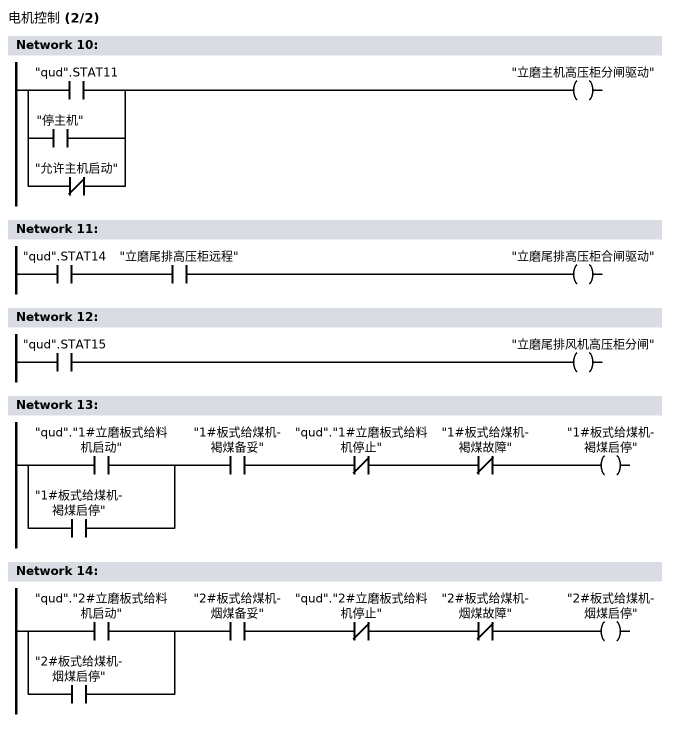
   RUNG wire#powerrail
      Contact( "qud".STAT11 )
      wire#w1
      Coil( "立磨主机高压柜分闸驱动" )
   END_RUNG
   RUNG wire#powerrail
      Contact( "停主机" )
   END_RUNG wire#w1
   RUNG wire#powerrail
      I_Contact( "允许主机启动" )
   END_RUNG wire#w1
   // the same network as SCL:
   "立磨主机高压柜分闸驱动" := "qud".STAT11 OR "停主机" OR NOT "允许主机启动";
END_REGION

REGION Network 11
   RUNG wire#powerrail
      Contact( "qud".STAT14 )
      Contact( "立磨尾排高压柜远程" )
      Coil( "立磨尾排高压柜合闸驱动" )
   END_RUNG
   // the same network as SCL:
   "立磨尾排高压柜合闸驱动" := "qud".STAT14 AND "立磨尾排高压柜远程";
END_REGION

REGION Network 12
   RUNG wire#powerrail
      Contact( "qud".STAT15 )
      Coil( "立磨尾排风机高压柜分闸" )
   END_RUNG
   // the same network as SCL:
   "立磨尾排风机高压柜分闸" := "qud".STAT15;
END_REGION

REGION Network 13
   RUNG wire#powerrail
      Contact( "qud"."1#立磨板式给料机启动" )
      wire#w1
      Contact( "1#板式给煤机-褐煤备妥" )
      I_Contact( "qud"."1#立磨板式给料机停止" )
      I_Contact( "1#板式给煤机-褐煤故障" )
      Coil( "1#板式给煤机-褐煤启停" )
   END_RUNG
   RUNG wire#powerrail
      Contact( "1#板式给煤机-褐煤启停" )
   END_RUNG wire#w1
   // the same network as SCL:
   "1#板式给煤机-褐煤启停" := ("qud"."1#立磨板式给料机启动" OR "1#板式给煤机-褐煤启停") AND "1#板式给煤机-褐煤备妥" AND NOT "qud"."1#立磨板式给料机停止" AND NOT "1#板式给煤机-褐煤故障";
END_REGION

REGION Network 14
   RUNG wire#powerrail
      Contact( "qud"."2#立磨板式给料机启动" )
      wire#w1
      Contact( "2#板式给煤机-烟煤备妥" )
      I_Contact( "qud"."2#立磨板式给料机停止" )
      I_Contact( "2#板式给煤机-烟煤故障" )
      Coil( "2#板式给煤机-烟煤启停" )
   END_RUNG
   RUNG wire#powerrail
      Contact( "2#板式给煤机-烟煤启停" )
   END_RUNG wire#w1
   // the same network as SCL:
   "2#板式给煤机-烟煤启停" := ("qud"."2#立磨板式给料机启动" OR "2#板式给煤机-烟煤启停") AND "2#板式给煤机-烟煤备妥" AND NOT "qud"."2#立磨板式给料机停止" AND NOT "2#板式给煤机-烟煤故障";
END_REGION
END_FUNCTION

FUNCTION "模拟量" : Void   // FC2, LAD
{ S7_Optimized_Access := 'FALSE' }
VERSION : 0.1
BEGIN

REGION Network 1
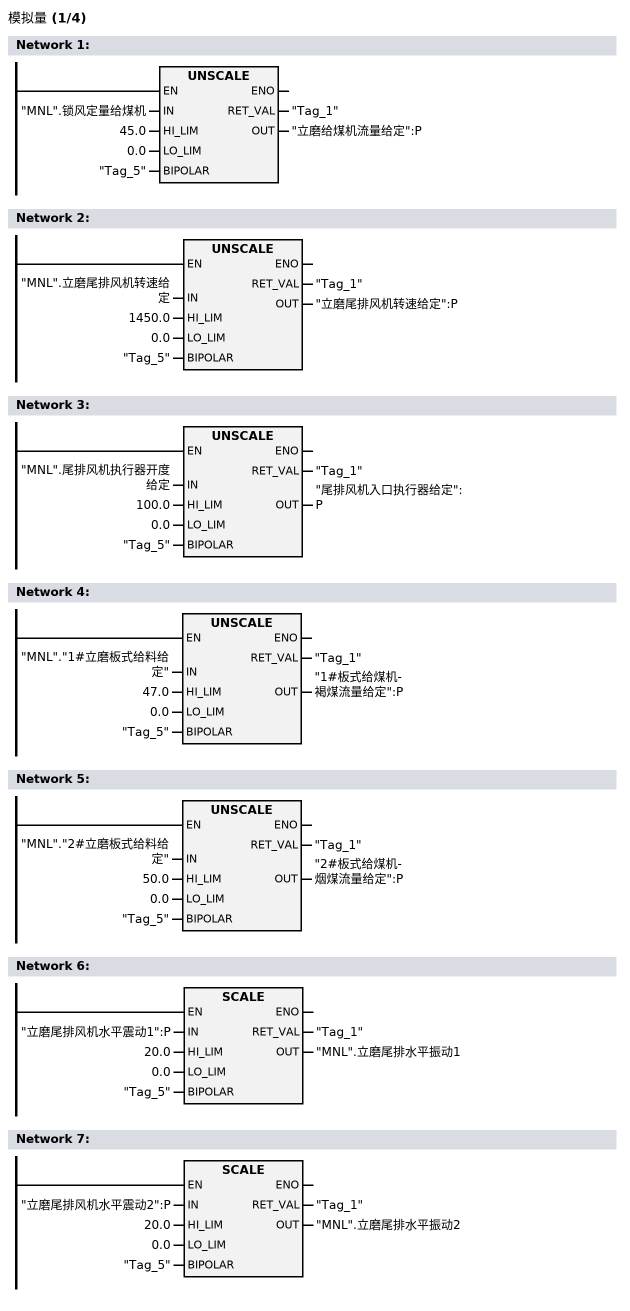
   "Tag_1" := UNSCALE(IN := "MNL".锁风定量给煤机,
                      HI_LIM := 45.0,
                      LO_LIM := 0.0,
                      BIPOLAR := "Tag_5",
                      OUT => "立磨给煤机流量给定":P);
END_REGION

REGION Network 2
   "Tag_1" := UNSCALE(IN := "MNL".立磨尾排风机转速给定,
                      HI_LIM := 1450.0,
                      LO_LIM := 0.0,
                      BIPOLAR := "Tag_5",
                      OUT => "立磨尾排风机转速给定":P);
END_REGION

REGION Network 3
   "Tag_1" := UNSCALE(IN := "MNL".尾排风机执行器开度给定,
                      HI_LIM := 100.0,
                      LO_LIM := 0.0,
                      BIPOLAR := "Tag_5",
                      OUT => "尾排风机入口执行器给定":P);
END_REGION

REGION Network 4
   "Tag_1" := UNSCALE(IN := "MNL"."1#立磨板式给料给定",
                      HI_LIM := 47.0,
                      LO_LIM := 0.0,
                      BIPOLAR := "Tag_5",
                      OUT => "1#板式给煤机-褐煤流量给定":P);
END_REGION

REGION Network 5
   "Tag_1" := UNSCALE(IN := "MNL"."2#立磨板式给料给定",
                      HI_LIM := 50.0,
                      LO_LIM := 0.0,
                      BIPOLAR := "Tag_5",
                      OUT => "2#板式给煤机-烟煤流量给定":P);
END_REGION

REGION Network 6
   "Tag_1" := SCALE(IN := "立磨尾排风机水平震动1":P,
                    HI_LIM := 20.0,
                    LO_LIM := 0.0,
                    BIPOLAR := "Tag_5",
                    OUT => "MNL".立磨尾排水平振动1);
END_REGION

REGION Network 7
   "Tag_1" := SCALE(IN := "立磨尾排风机水平震动2":P,
                    HI_LIM := 20.0,
                    LO_LIM := 0.0,
                    BIPOLAR := "Tag_5",
                    OUT => "MNL".立磨尾排水平振动2);
END_REGION

REGION Network 8
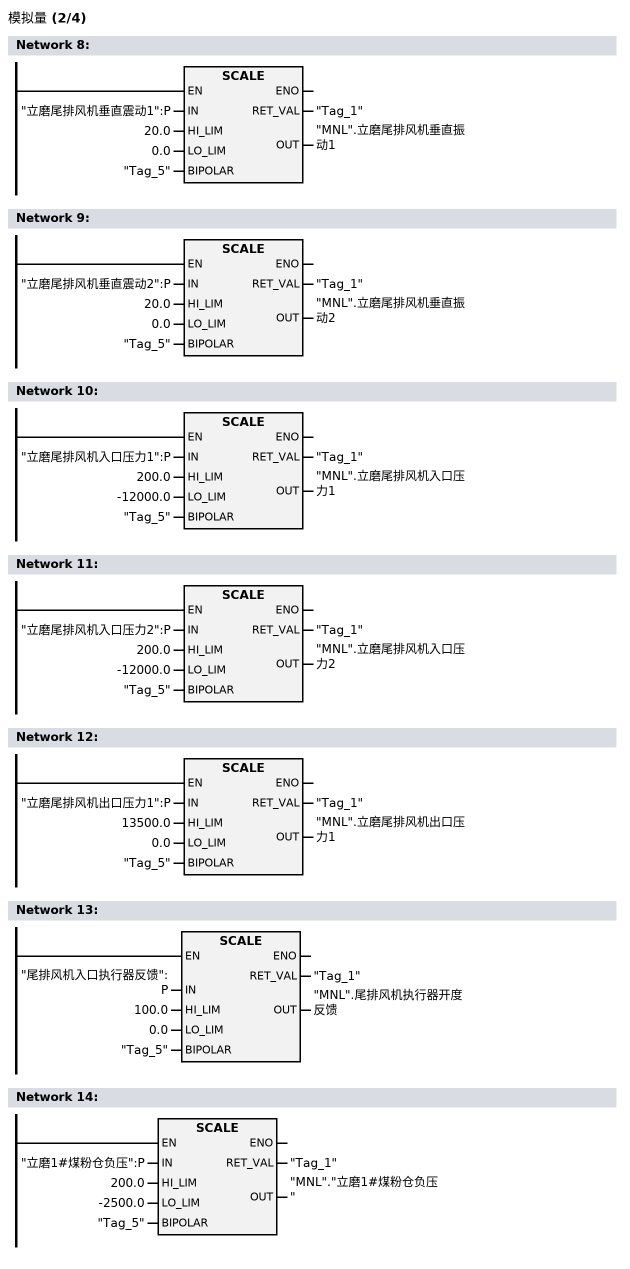
   "Tag_1" := SCALE(IN := "立磨尾排风机垂直震动1":P,
                    HI_LIM := 20.0,
                    LO_LIM := 0.0,
                    BIPOLAR := "Tag_5",
                    OUT => "MNL".立磨尾排风机垂直振动1);
END_REGION

REGION Network 9
   "Tag_1" := SCALE(IN := "立磨尾排风机垂直震动2":P,
                    HI_LIM := 20.0,
                    LO_LIM := 0.0,
                    BIPOLAR := "Tag_5",
                    OUT => "MNL".立磨尾排风机垂直振动2);
END_REGION

REGION Network 10
   "Tag_1" := SCALE(IN := "立磨尾排风机入口压力1":P,
                    HI_LIM := 200.0,
                    LO_LIM := -12000.0,
                    BIPOLAR := "Tag_5",
                    OUT => "MNL".立磨尾排风机入口压力1);
END_REGION

REGION Network 11
   "Tag_1" := SCALE(IN := "立磨尾排风机入口压力2":P,
                    HI_LIM := 200.0,
                    LO_LIM := -12000.0,
                    BIPOLAR := "Tag_5",
                    OUT => "MNL".立磨尾排风机入口压力2);
END_REGION

REGION Network 12
   "Tag_1" := SCALE(IN := "立磨尾排风机出口压力1":P,
                    HI_LIM := 13500.0,
                    LO_LIM := 0.0,
                    BIPOLAR := "Tag_5",
                    OUT => "MNL".立磨尾排风机出口压力1);
END_REGION

REGION Network 13
   "Tag_1" := SCALE(IN := "尾排风机入口执行器反馈":P,
                    HI_LIM := 100.0,
                    LO_LIM := 0.0,
                    BIPOLAR := "Tag_5",
                    OUT => "MNL".尾排风机执行器开度反馈);
END_REGION

REGION Network 14
   "Tag_1" := SCALE(IN := "立磨1#煤粉仓负压":P,
                    HI_LIM := 200.0,
                    LO_LIM := -2500.0,
                    BIPOLAR := "Tag_5",
                    OUT => "MNL"."立磨1#煤粉仓负压");
END_REGION

REGION Network 15
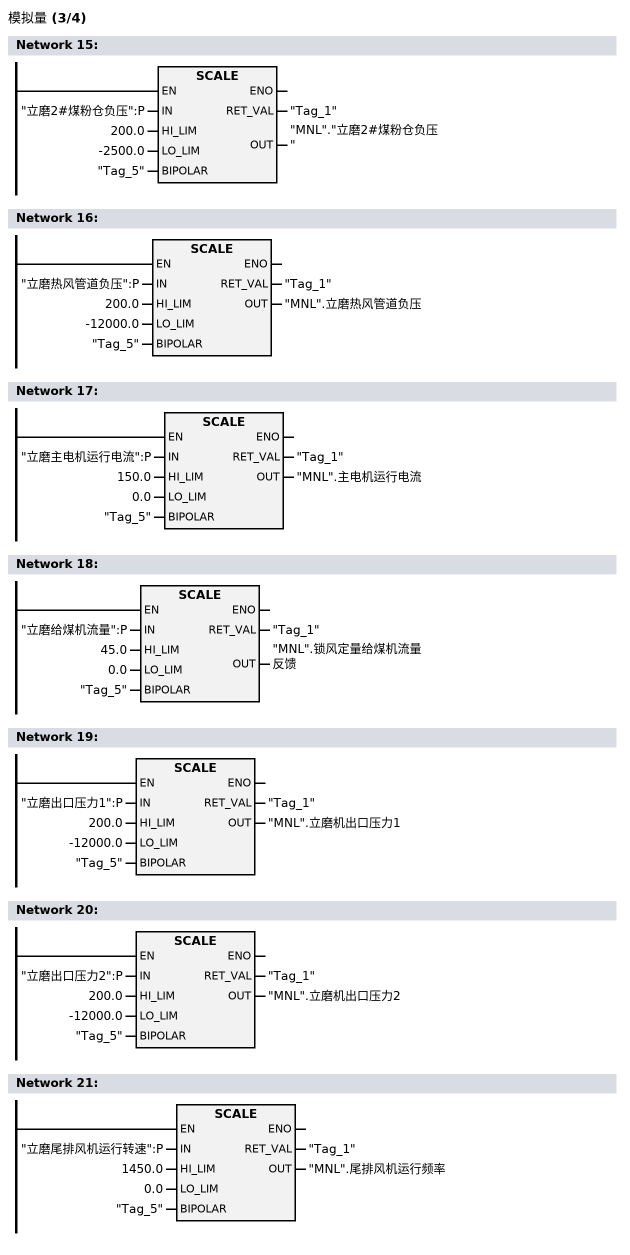
   "Tag_1" := SCALE(IN := "立磨2#煤粉仓负压":P,
                    HI_LIM := 200.0,
                    LO_LIM := -2500.0,
                    BIPOLAR := "Tag_5",
                    OUT => "MNL"."立磨2#煤粉仓负压");
END_REGION

REGION Network 16
   "Tag_1" := SCALE(IN := "立磨热风管道负压":P,
                    HI_LIM := 200.0,
                    LO_LIM := -12000.0,
                    BIPOLAR := "Tag_5",
                    OUT => "MNL".立磨热风管道负压);
END_REGION

REGION Network 17
   "Tag_1" := SCALE(IN := "立磨主电机运行电流":P,
                    HI_LIM := 150.0,
                    LO_LIM := 0.0,
                    BIPOLAR := "Tag_5",
                    OUT => "MNL".主电机运行电流);
END_REGION

REGION Network 18
   "Tag_1" := SCALE(IN := "立磨给煤机流量":P,
                    HI_LIM := 45.0,
                    LO_LIM := 0.0,
                    BIPOLAR := "Tag_5",
                    OUT => "MNL".锁风定量给煤机流量反馈);
END_REGION

REGION Network 19
   "Tag_1" := SCALE(IN := "立磨出口压力1":P,
                    HI_LIM := 200.0,
                    LO_LIM := -12000.0,
                    BIPOLAR := "Tag_5",
                    OUT => "MNL".立磨机出口压力1);
END_REGION

REGION Network 20
   "Tag_1" := SCALE(IN := "立磨出口压力2":P,
                    HI_LIM := 200.0,
                    LO_LIM := -12000.0,
                    BIPOLAR := "Tag_5",
                    OUT => "MNL".立磨机出口压力2);
END_REGION

REGION Network 21
   "Tag_1" := SCALE(IN := "立磨尾排风机运行转速":P,
                    HI_LIM := 1450.0,
                    LO_LIM := 0.0,
                    BIPOLAR := "Tag_5",
                    OUT => "MNL".尾排风机运行频率);
END_REGION

REGION Network 22
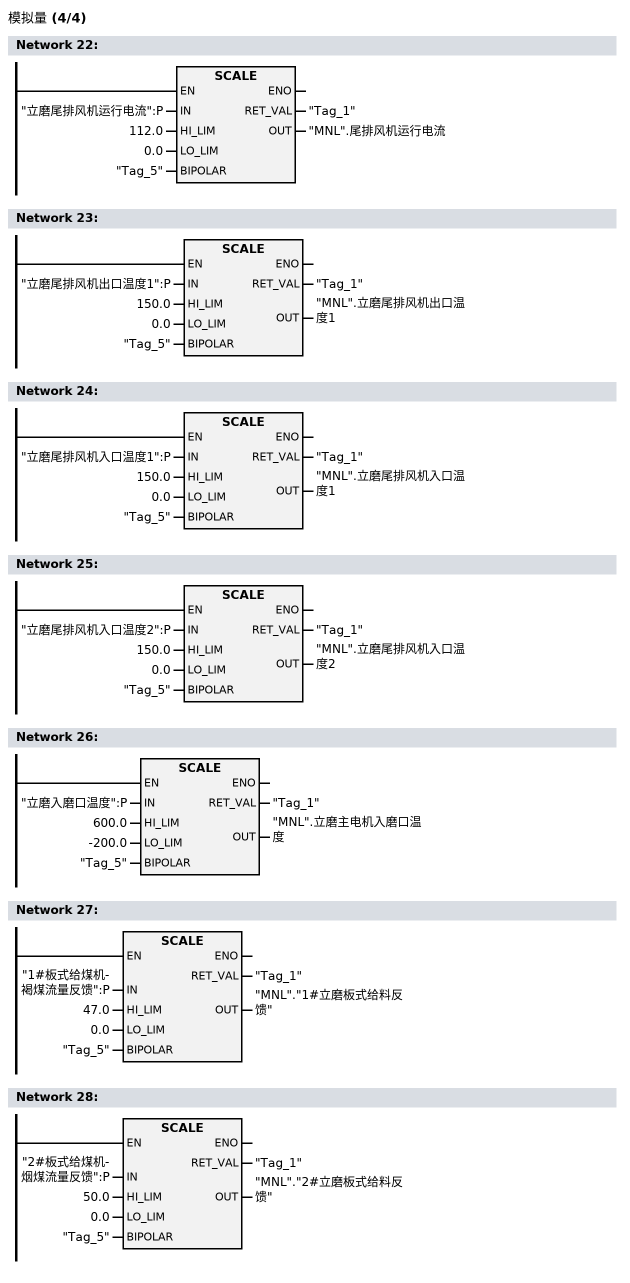
   "Tag_1" := SCALE(IN := "立磨尾排风机运行电流":P,
                    HI_LIM := 112.0,
                    LO_LIM := 0.0,
                    BIPOLAR := "Tag_5",
                    OUT => "MNL".尾排风机运行电流);
END_REGION

REGION Network 23
   "Tag_1" := SCALE(IN := "立磨尾排风机出口温度1":P,
                    HI_LIM := 150.0,
                    LO_LIM := 0.0,
                    BIPOLAR := "Tag_5",
                    OUT => "MNL".立磨尾排风机出口温度1);
END_REGION

REGION Network 24
   "Tag_1" := SCALE(IN := "立磨尾排风机入口温度1":P,
                    HI_LIM := 150.0,
                    LO_LIM := 0.0,
                    BIPOLAR := "Tag_5",
                    OUT => "MNL".立磨尾排风机入口温度1);
END_REGION

REGION Network 25
   "Tag_1" := SCALE(IN := "立磨尾排风机入口温度2":P,
                    HI_LIM := 150.0,
                    LO_LIM := 0.0,
                    BIPOLAR := "Tag_5",
                    OUT => "MNL".立磨尾排风机入口温度2);
END_REGION

REGION Network 26
   "Tag_1" := SCALE(IN := "立磨入磨口温度":P,
                    HI_LIM := 600.0,
                    LO_LIM := -200.0,
                    BIPOLAR := "Tag_5",
                    OUT => "MNL".立磨主电机入磨口温度);
END_REGION

REGION Network 27
   "Tag_1" := SCALE(IN := "1#板式给煤机-褐煤流量反馈":P,
                    HI_LIM := 47.0,
                    LO_LIM := 0.0,
                    BIPOLAR := "Tag_5",
                    OUT => "MNL"."1#立磨板式给料反馈");
END_REGION

REGION Network 28
   "Tag_1" := SCALE(IN := "2#板式给煤机-烟煤流量反馈":P,
                    HI_LIM := 50.0,
                    LO_LIM := 0.0,
                    BIPOLAR := "Tag_5",
                    OUT => "MNL"."2#立磨板式给料反馈");
END_REGION
END_FUNCTION

FUNCTION "料仓控制" : Void   // FC3, LAD
{ S7_Optimized_Access := 'FALSE' }
VERSION : 0.1
BEGIN

REGION Network 1
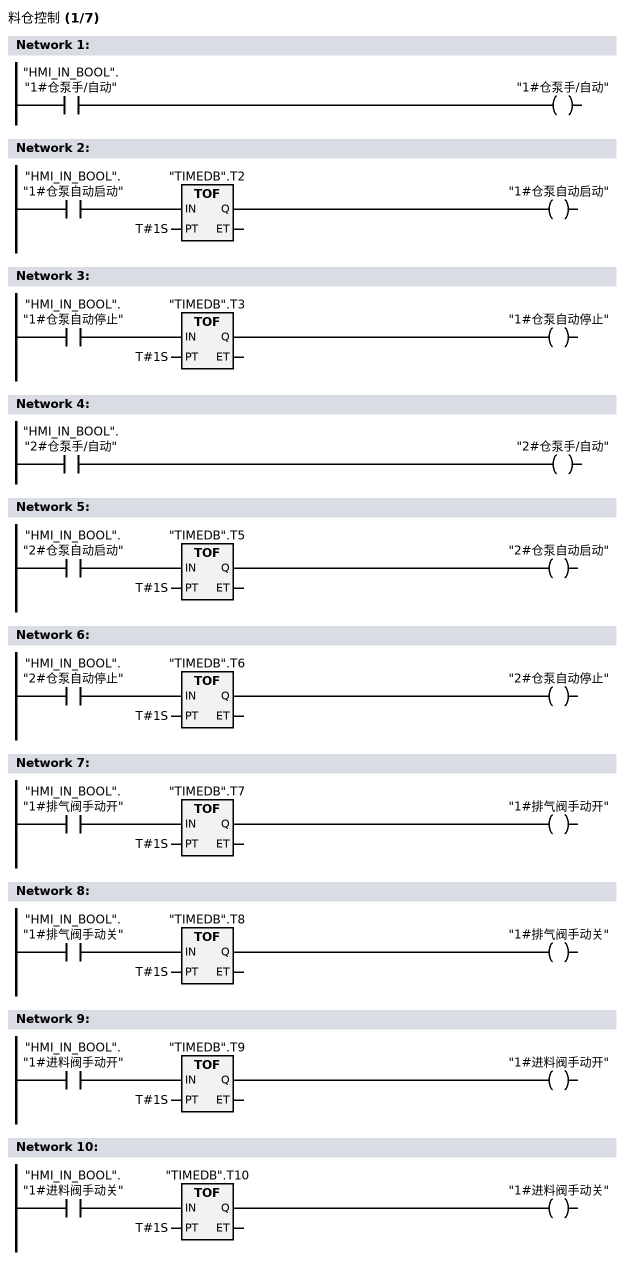
   RUNG wire#powerrail
      Contact( "HMI_IN_BOOL"."1#仓泵手/自动" )
      Coil( "1#仓泵手/自动" )
   END_RUNG
   // the same network as SCL:
   "1#仓泵手/自动" := "HMI_IN_BOOL"."1#仓泵手/自动";
END_REGION

REGION Network 2
   "TIMEDB".T2.TOF(IN := "HMI_IN_BOOL"."1#仓泵自动启动", PT := T#1S);
   "1#仓泵自动启动" := "TIMEDB".T2.Q;
END_REGION

REGION Network 3
   "TIMEDB".T3.TOF(IN := "HMI_IN_BOOL"."1#仓泵自动停止", PT := T#1S);
   "1#仓泵自动停止" := "TIMEDB".T3.Q;
END_REGION

REGION Network 4
   RUNG wire#powerrail
      Contact( "HMI_IN_BOOL"."2#仓泵手/自动" )
      Coil( "2#仓泵手/自动" )
   END_RUNG
   // the same network as SCL:
   "2#仓泵手/自动" := "HMI_IN_BOOL"."2#仓泵手/自动";
END_REGION

REGION Network 5
   "TIMEDB".T5.TOF(IN := "HMI_IN_BOOL"."2#仓泵自动启动", PT := T#1S);
   "2#仓泵自动启动" := "TIMEDB".T5.Q;
END_REGION

REGION Network 6
   "TIMEDB".T6.TOF(IN := "HMI_IN_BOOL"."2#仓泵自动停止", PT := T#1S);
   "2#仓泵自动停止" := "TIMEDB".T6.Q;
END_REGION

REGION Network 7
   "TIMEDB".T7.TOF(IN := "HMI_IN_BOOL"."1#排气阀手动开", PT := T#1S);
   "1#排气阀手动开" := "TIMEDB".T7.Q;
END_REGION

REGION Network 8
   "TIMEDB".T8.TOF(IN := "HMI_IN_BOOL"."1#排气阀手动关", PT := T#1S);
   "1#排气阀手动关" := "TIMEDB".T8.Q;
END_REGION

REGION Network 9
   "TIMEDB".T9.TOF(IN := "HMI_IN_BOOL"."1#进料阀手动开", PT := T#1S);
   "1#进料阀手动开" := "TIMEDB".T9.Q;
END_REGION

REGION Network 10
   "TIMEDB".T10.TOF(IN := "HMI_IN_BOOL"."1#进料阀手动关", PT := T#1S);
   "1#进料阀手动关" := "TIMEDB".T10.Q;
END_REGION

REGION Network 11
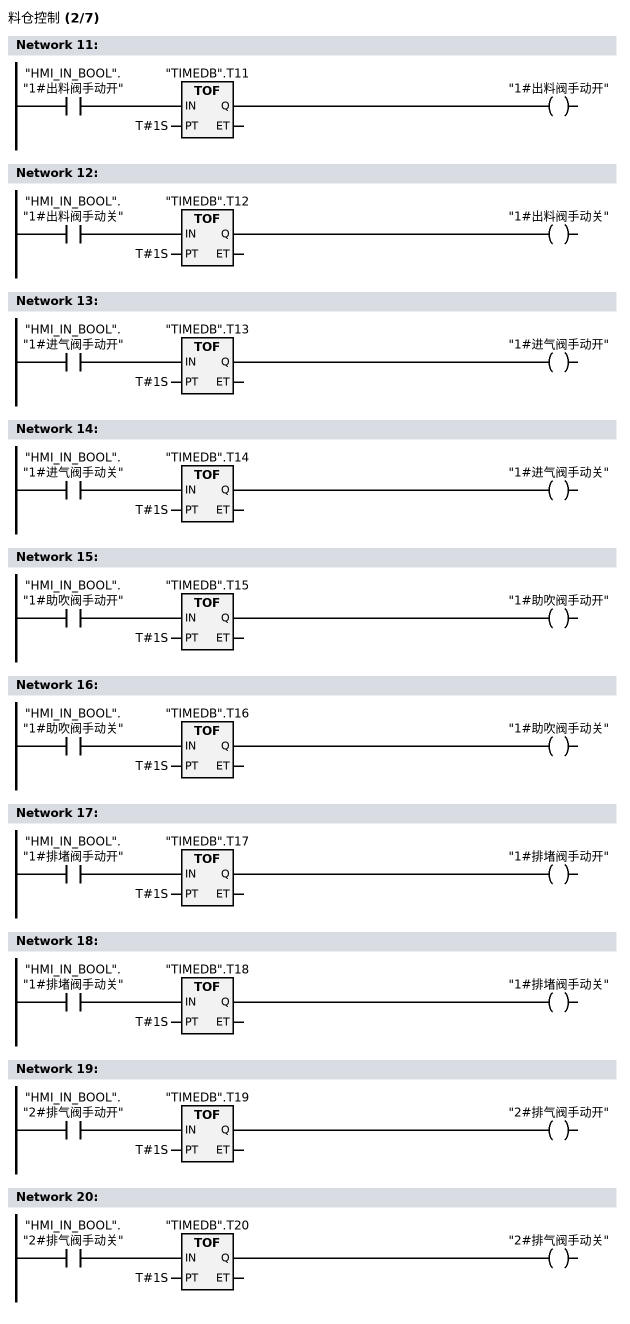
   "TIMEDB".T11.TOF(IN := "HMI_IN_BOOL"."1#出料阀手动开", PT := T#1S);
   "1#出料阀手动开" := "TIMEDB".T11.Q;
END_REGION

REGION Network 12
   "TIMEDB".T12.TOF(IN := "HMI_IN_BOOL"."1#出料阀手动关", PT := T#1S);
   "1#出料阀手动关" := "TIMEDB".T12.Q;
END_REGION

REGION Network 13
   "TIMEDB".T13.TOF(IN := "HMI_IN_BOOL"."1#进气阀手动开", PT := T#1S);
   "1#进气阀手动开" := "TIMEDB".T13.Q;
END_REGION

REGION Network 14
   "TIMEDB".T14.TOF(IN := "HMI_IN_BOOL"."1#进气阀手动关", PT := T#1S);
   "1#进气阀手动关" := "TIMEDB".T14.Q;
END_REGION

REGION Network 15
   "TIMEDB".T15.TOF(IN := "HMI_IN_BOOL"."1#助吹阀手动开", PT := T#1S);
   "1#助吹阀手动开" := "TIMEDB".T15.Q;
END_REGION

REGION Network 16
   "TIMEDB".T16.TOF(IN := "HMI_IN_BOOL"."1#助吹阀手动关", PT := T#1S);
   "1#助吹阀手动关" := "TIMEDB".T16.Q;
END_REGION

REGION Network 17
   "TIMEDB".T17.TOF(IN := "HMI_IN_BOOL"."1#排堵阀手动开", PT := T#1S);
   "1#排堵阀手动开" := "TIMEDB".T17.Q;
END_REGION

REGION Network 18
   "TIMEDB".T18.TOF(IN := "HMI_IN_BOOL"."1#排堵阀手动关", PT := T#1S);
   "1#排堵阀手动关" := "TIMEDB".T18.Q;
END_REGION

REGION Network 19
   "TIMEDB".T19.TOF(IN := "HMI_IN_BOOL"."2#排气阀手动开", PT := T#1S);
   "2#排气阀手动开" := "TIMEDB".T19.Q;
END_REGION

REGION Network 20
   "TIMEDB".T20.TOF(IN := "HMI_IN_BOOL"."2#排气阀手动关", PT := T#1S);
   "2#排气阀手动关" := "TIMEDB".T20.Q;
END_REGION

REGION Network 21
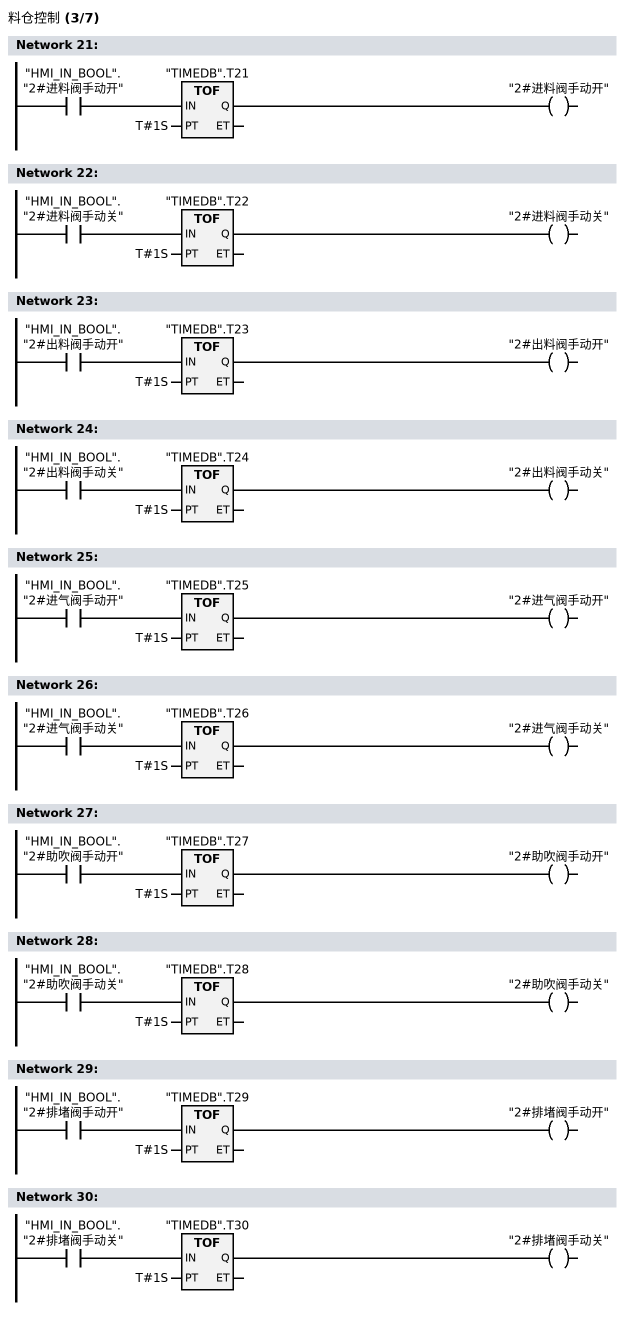
   "TIMEDB".T21.TOF(IN := "HMI_IN_BOOL"."2#进料阀手动开", PT := T#1S);
   "2#进料阀手动开" := "TIMEDB".T21.Q;
END_REGION

REGION Network 22
   "TIMEDB".T22.TOF(IN := "HMI_IN_BOOL"."2#进料阀手动关", PT := T#1S);
   "2#进料阀手动关" := "TIMEDB".T22.Q;
END_REGION

REGION Network 23
   "TIMEDB".T23.TOF(IN := "HMI_IN_BOOL"."2#出料阀手动开", PT := T#1S);
   "2#出料阀手动开" := "TIMEDB".T23.Q;
END_REGION

REGION Network 24
   "TIMEDB".T24.TOF(IN := "HMI_IN_BOOL"."2#出料阀手动关", PT := T#1S);
   "2#出料阀手动关" := "TIMEDB".T24.Q;
END_REGION

REGION Network 25
   "TIMEDB".T25.TOF(IN := "HMI_IN_BOOL"."2#进气阀手动开", PT := T#1S);
   "2#进气阀手动开" := "TIMEDB".T25.Q;
END_REGION

REGION Network 26
   "TIMEDB".T26.TOF(IN := "HMI_IN_BOOL"."2#进气阀手动关", PT := T#1S);
   "2#进气阀手动关" := "TIMEDB".T26.Q;
END_REGION

REGION Network 27
   "TIMEDB".T27.TOF(IN := "HMI_IN_BOOL"."2#助吹阀手动开", PT := T#1S);
   "2#助吹阀手动开" := "TIMEDB".T27.Q;
END_REGION

REGION Network 28
   "TIMEDB".T28.TOF(IN := "HMI_IN_BOOL"."2#助吹阀手动关", PT := T#1S);
   "2#助吹阀手动关" := "TIMEDB".T28.Q;
END_REGION

REGION Network 29
   "TIMEDB".T29.TOF(IN := "HMI_IN_BOOL"."2#排堵阀手动开", PT := T#1S);
   "2#排堵阀手动开" := "TIMEDB".T29.Q;
END_REGION

REGION Network 30
   "TIMEDB".T30.TOF(IN := "HMI_IN_BOOL"."2#排堵阀手动关", PT := T#1S);
   "2#排堵阀手动关" := "TIMEDB".T30.Q;
END_REGION

REGION Network 31
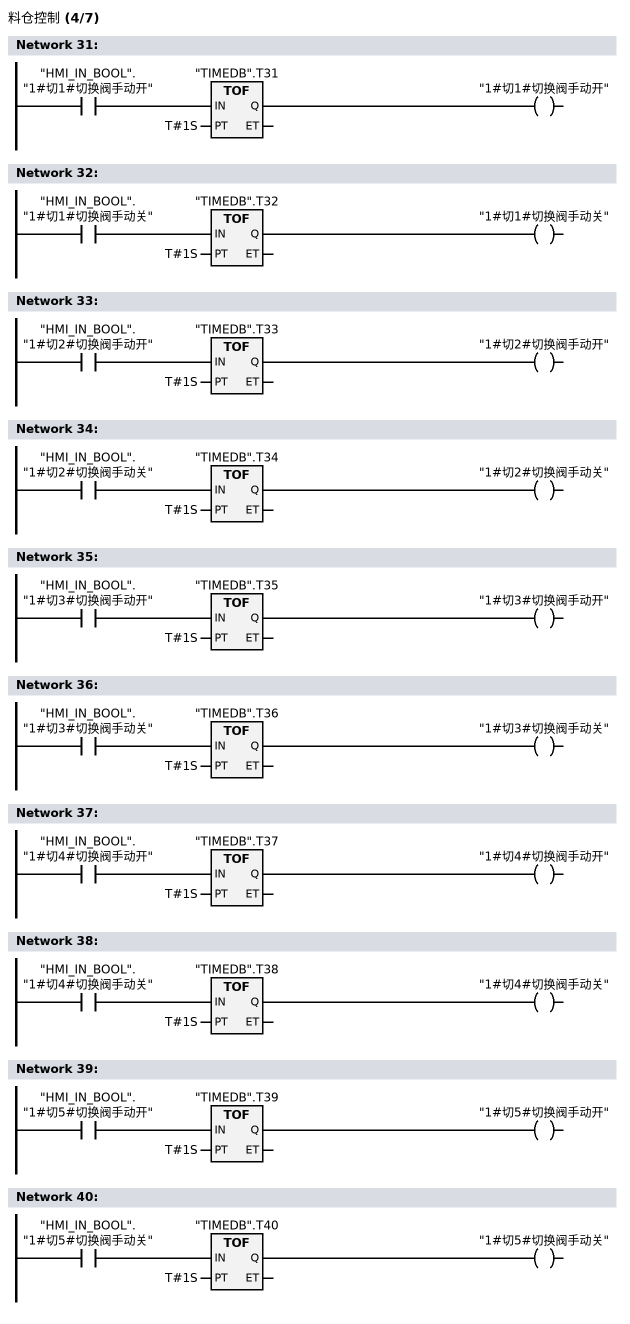
   "TIMEDB".T31.TOF(IN := "HMI_IN_BOOL"."1#切1#切换阀手动开", PT := T#1S);
   "1#切1#切换阀手动开" := "TIMEDB".T31.Q;
END_REGION

REGION Network 32
   "TIMEDB".T32.TOF(IN := "HMI_IN_BOOL"."1#切1#切换阀手动关", PT := T#1S);
   "1#切1#切换阀手动关" := "TIMEDB".T32.Q;
END_REGION

REGION Network 33
   "TIMEDB".T33.TOF(IN := "HMI_IN_BOOL"."1#切2#切换阀手动开", PT := T#1S);
   "1#切2#切换阀手动开" := "TIMEDB".T33.Q;
END_REGION

REGION Network 34
   "TIMEDB".T34.TOF(IN := "HMI_IN_BOOL"."1#切2#切换阀手动关", PT := T#1S);
   "1#切2#切换阀手动关" := "TIMEDB".T34.Q;
END_REGION

REGION Network 35
   "TIMEDB".T35.TOF(IN := "HMI_IN_BOOL"."1#切3#切换阀手动开", PT := T#1S);
   "1#切3#切换阀手动开" := "TIMEDB".T35.Q;
END_REGION

REGION Network 36
   "TIMEDB".T36.TOF(IN := "HMI_IN_BOOL"."1#切3#切换阀手动关", PT := T#1S);
   "1#切3#切换阀手动关" := "TIMEDB".T36.Q;
END_REGION

REGION Network 37
   "TIMEDB".T37.TOF(IN := "HMI_IN_BOOL"."1#切4#切换阀手动开", PT := T#1S);
   "1#切4#切换阀手动开" := "TIMEDB".T37.Q;
END_REGION

REGION Network 38
   "TIMEDB".T38.TOF(IN := "HMI_IN_BOOL"."1#切4#切换阀手动关", PT := T#1S);
   "1#切4#切换阀手动关" := "TIMEDB".T38.Q;
END_REGION

REGION Network 39
   "TIMEDB".T39.TOF(IN := "HMI_IN_BOOL"."1#切5#切换阀手动开", PT := T#1S);
   "1#切5#切换阀手动开" := "TIMEDB".T39.Q;
END_REGION

REGION Network 40
   "TIMEDB".T40.TOF(IN := "HMI_IN_BOOL"."1#切5#切换阀手动关", PT := T#1S);
   "1#切5#切换阀手动关" := "TIMEDB".T40.Q;
END_REGION

REGION Network 41
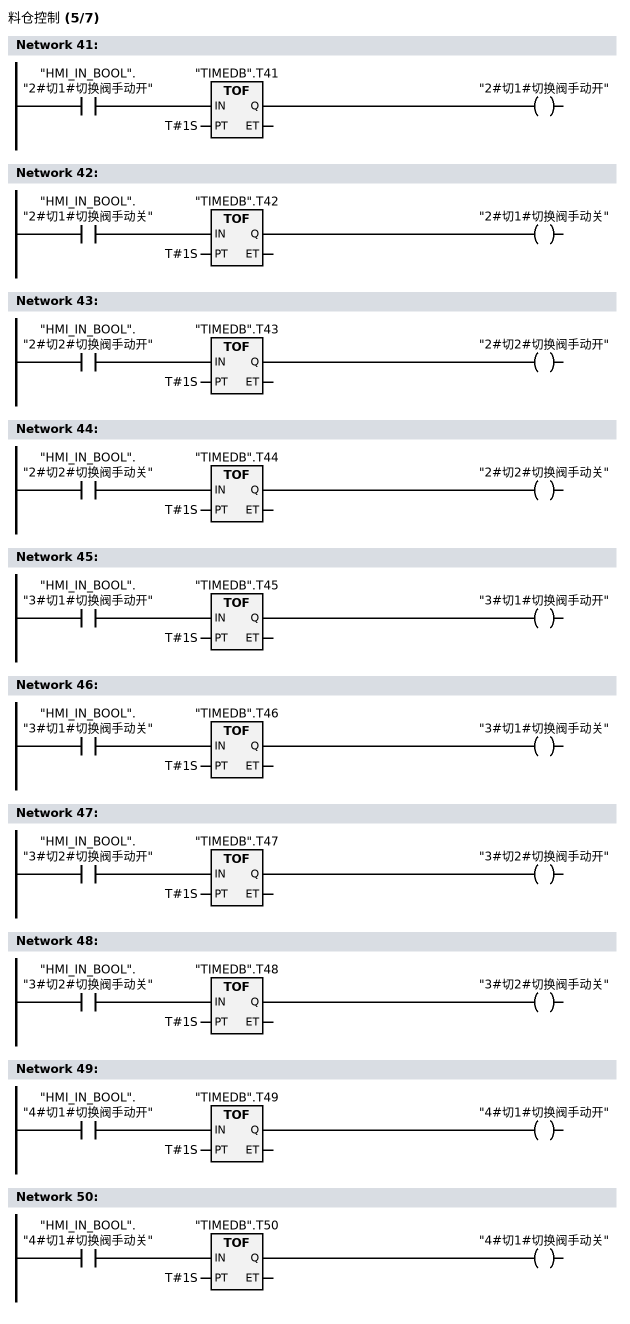
   "TIMEDB".T41.TOF(IN := "HMI_IN_BOOL"."2#切1#切换阀手动开", PT := T#1S);
   "2#切1#切换阀手动开" := "TIMEDB".T41.Q;
END_REGION

REGION Network 42
   "TIMEDB".T42.TOF(IN := "HMI_IN_BOOL"."2#切1#切换阀手动关", PT := T#1S);
   "2#切1#切换阀手动关" := "TIMEDB".T42.Q;
END_REGION

REGION Network 43
   "TIMEDB".T43.TOF(IN := "HMI_IN_BOOL"."2#切2#切换阀手动开", PT := T#1S);
   "2#切2#切换阀手动开" := "TIMEDB".T43.Q;
END_REGION

REGION Network 44
   "TIMEDB".T44.TOF(IN := "HMI_IN_BOOL"."2#切2#切换阀手动关", PT := T#1S);
   "2#切2#切换阀手动关" := "TIMEDB".T44.Q;
END_REGION

REGION Network 45
   "TIMEDB".T45.TOF(IN := "HMI_IN_BOOL"."3#切1#切换阀手动开", PT := T#1S);
   "3#切1#切换阀手动开" := "TIMEDB".T45.Q;
END_REGION

REGION Network 46
   "TIMEDB".T46.TOF(IN := "HMI_IN_BOOL"."3#切1#切换阀手动关", PT := T#1S);
   "3#切1#切换阀手动关" := "TIMEDB".T46.Q;
END_REGION

REGION Network 47
   "TIMEDB".T47.TOF(IN := "HMI_IN_BOOL"."3#切2#切换阀手动开", PT := T#1S);
   "3#切2#切换阀手动开" := "TIMEDB".T47.Q;
END_REGION

REGION Network 48
   "TIMEDB".T48.TOF(IN := "HMI_IN_BOOL"."3#切2#切换阀手动关", PT := T#1S);
   "3#切2#切换阀手动关" := "TIMEDB".T48.Q;
END_REGION

REGION Network 49
   "TIMEDB".T49.TOF(IN := "HMI_IN_BOOL"."4#切1#切换阀手动开", PT := T#1S);
   "4#切1#切换阀手动开" := "TIMEDB".T49.Q;
END_REGION

REGION Network 50
   "TIMEDB".T50.TOF(IN := "HMI_IN_BOOL"."4#切1#切换阀手动关", PT := T#1S);
   "4#切1#切换阀手动关" := "TIMEDB".T50.Q;
END_REGION

REGION Network 51
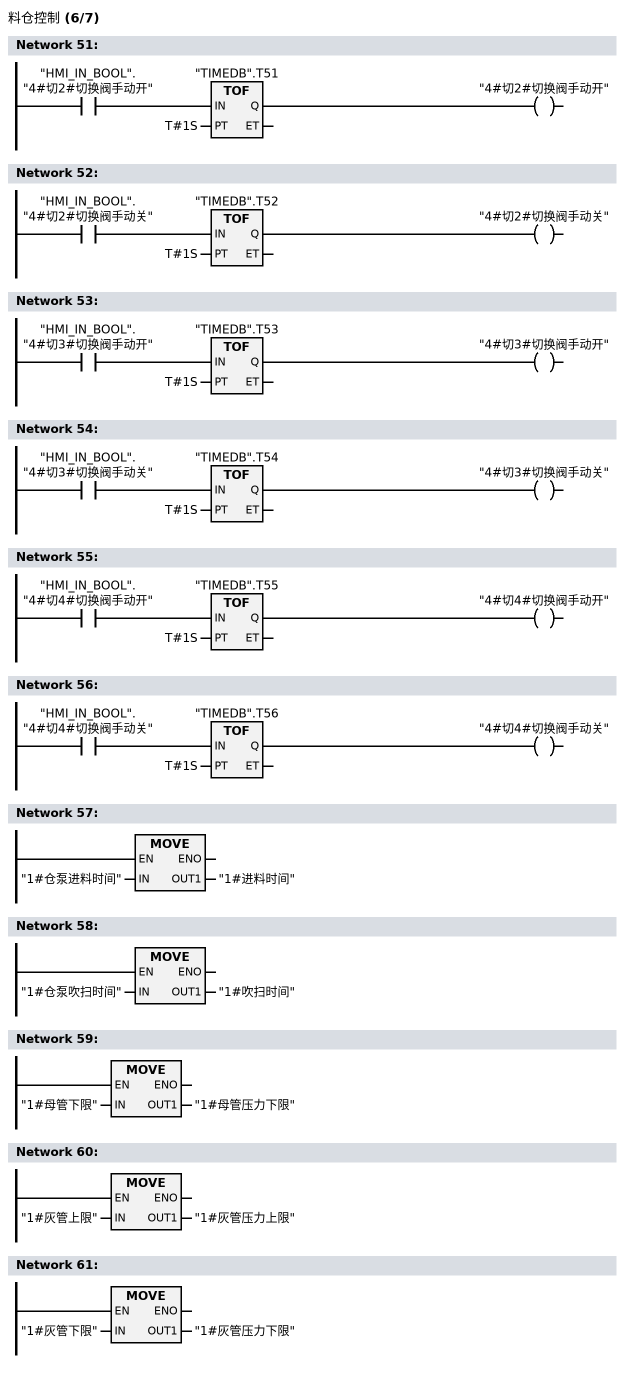
   "TIMEDB".T51.TOF(IN := "HMI_IN_BOOL"."4#切2#切换阀手动开", PT := T#1S);
   "4#切2#切换阀手动开" := "TIMEDB".T51.Q;
END_REGION

REGION Network 52
   "TIMEDB".T52.TOF(IN := "HMI_IN_BOOL"."4#切2#切换阀手动关", PT := T#1S);
   "4#切2#切换阀手动关" := "TIMEDB".T52.Q;
END_REGION

REGION Network 53
   "TIMEDB".T53.TOF(IN := "HMI_IN_BOOL"."4#切3#切换阀手动开", PT := T#1S);
   "4#切3#切换阀手动开" := "TIMEDB".T53.Q;
END_REGION

REGION Network 54
   "TIMEDB".T54.TOF(IN := "HMI_IN_BOOL"."4#切3#切换阀手动关", PT := T#1S);
   "4#切3#切换阀手动关" := "TIMEDB".T54.Q;
END_REGION

REGION Network 55
   "TIMEDB".T55.TOF(IN := "HMI_IN_BOOL"."4#切4#切换阀手动开", PT := T#1S);
   "4#切4#切换阀手动开" := "TIMEDB".T55.Q;
END_REGION

REGION Network 56
   "TIMEDB".T56.TOF(IN := "HMI_IN_BOOL"."4#切4#切换阀手动关", PT := T#1S);
   "4#切4#切换阀手动关" := "TIMEDB".T56.Q;
END_REGION

REGION Network 57
   RUNG wire#powerrail
      { S7_GenerateENO := "TRUE" } Move(in := "1#仓泵进料时间", out1 => "1#进料时间")
   END_RUNG
   // the same network as SCL:
   "1#进料时间" := "1#仓泵进料时间";
END_REGION

REGION Network 58
   RUNG wire#powerrail
      { S7_GenerateENO := "TRUE" } Move(in := "1#仓泵吹扫时间", out1 => "1#吹扫时间")
   END_RUNG
   // the same network as SCL:
   "1#吹扫时间" := "1#仓泵吹扫时间";
END_REGION

REGION Network 59
   RUNG wire#powerrail
      { S7_GenerateENO := "TRUE" } Move(in := "1#母管下限", out1 => "1#母管压力下限")
   END_RUNG
   // the same network as SCL:
   "1#母管压力下限" := "1#母管下限";
END_REGION

REGION Network 60
   RUNG wire#powerrail
      { S7_GenerateENO := "TRUE" } Move(in := "1#灰管上限", out1 => "1#灰管压力上限")
   END_RUNG
   // the same network as SCL:
   "1#灰管压力上限" := "1#灰管上限";
END_REGION

REGION Network 61
   RUNG wire#powerrail
      { S7_GenerateENO := "TRUE" } Move(in := "1#灰管下限", out1 => "1#灰管压力下限")
   END_RUNG
   // the same network as SCL:
   "1#灰管压力下限" := "1#灰管下限";
END_REGION

REGION Network 62
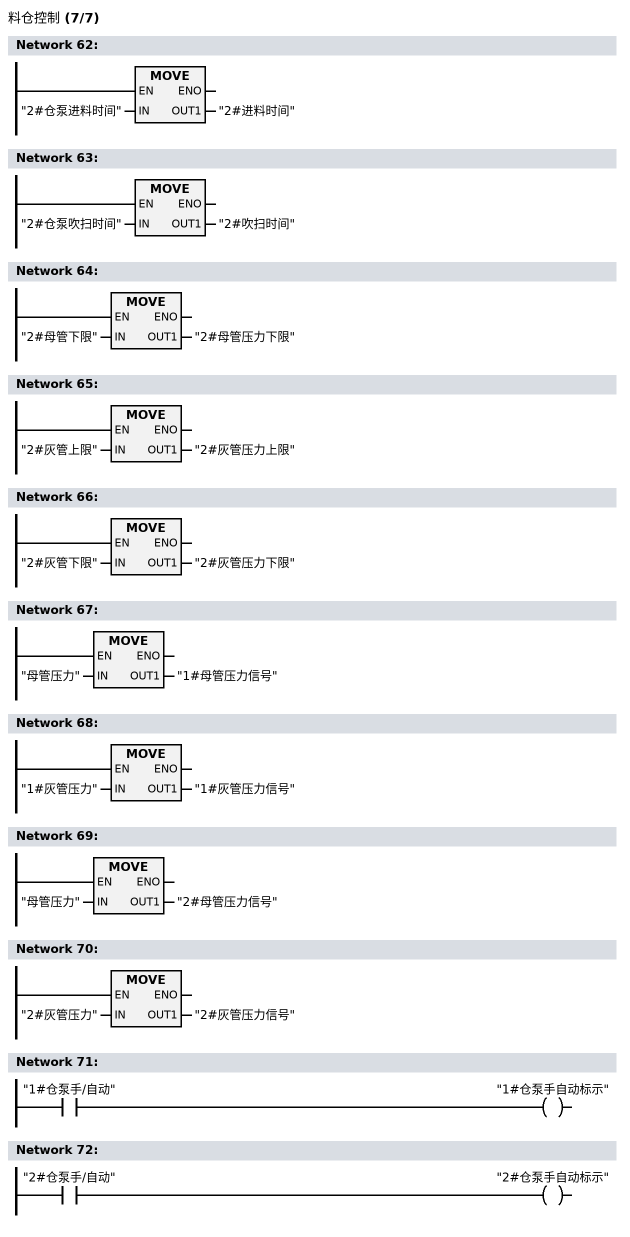
   RUNG wire#powerrail
      { S7_GenerateENO := "TRUE" } Move(in := "2#仓泵进料时间", out1 => "2#进料时间")
   END_RUNG
   // the same network as SCL:
   "2#进料时间" := "2#仓泵进料时间";
END_REGION

REGION Network 63
   RUNG wire#powerrail
      { S7_GenerateENO := "TRUE" } Move(in := "2#仓泵吹扫时间", out1 => "2#吹扫时间")
   END_RUNG
   // the same network as SCL:
   "2#吹扫时间" := "2#仓泵吹扫时间";
END_REGION

REGION Network 64
   RUNG wire#powerrail
      { S7_GenerateENO := "TRUE" } Move(in := "2#母管下限", out1 => "2#母管压力下限")
   END_RUNG
   // the same network as SCL:
   "2#母管压力下限" := "2#母管下限";
END_REGION

REGION Network 65
   RUNG wire#powerrail
      { S7_GenerateENO := "TRUE" } Move(in := "2#灰管上限", out1 => "2#灰管压力上限")
   END_RUNG
   // the same network as SCL:
   "2#灰管压力上限" := "2#灰管上限";
END_REGION

REGION Network 66
   RUNG wire#powerrail
      { S7_GenerateENO := "TRUE" } Move(in := "2#灰管下限", out1 => "2#灰管压力下限")
   END_RUNG
   // the same network as SCL:
   "2#灰管压力下限" := "2#灰管下限";
END_REGION

REGION Network 67
   RUNG wire#powerrail
      { S7_GenerateENO := "TRUE" } Move(in := "母管压力", out1 => "1#母管压力信号")
   END_RUNG
   // the same network as SCL:
   "1#母管压力信号" := "母管压力";
END_REGION

REGION Network 68
   RUNG wire#powerrail
      { S7_GenerateENO := "TRUE" } Move(in := "1#灰管压力", out1 => "1#灰管压力信号")
   END_RUNG
   // the same network as SCL:
   "1#灰管压力信号" := "1#灰管压力";
END_REGION

REGION Network 69
   RUNG wire#powerrail
      { S7_GenerateENO := "TRUE" } Move(in := "母管压力", out1 => "2#母管压力信号")
   END_RUNG
   // the same network as SCL:
   "2#母管压力信号" := "母管压力";
END_REGION

REGION Network 70
   RUNG wire#powerrail
      { S7_GenerateENO := "TRUE" } Move(in := "2#灰管压力", out1 => "2#灰管压力信号")
   END_RUNG
   // the same network as SCL:
   "2#灰管压力信号" := "2#灰管压力";
END_REGION

REGION Network 71
   RUNG wire#powerrail
      Contact( "1#仓泵手/自动" )
      Coil( "1#仓泵手自动标示" )
   END_RUNG
   // the same network as SCL:
   "1#仓泵手自动标示" := "1#仓泵手/自动";
END_REGION

REGION Network 72
   RUNG wire#powerrail
      Contact( "2#仓泵手/自动" )
      Coil( "2#仓泵手自动标示" )
   END_RUNG
   // the same network as SCL:
   "2#仓泵手自动标示" := "2#仓泵手/自动";
END_REGION
END_FUNCTION

FUNCTION "仪表数据" : Void   // FC4, LAD
{ S7_Optimized_Access := 'FALSE' }
VERSION : 0.1
BEGIN

REGION Network 1
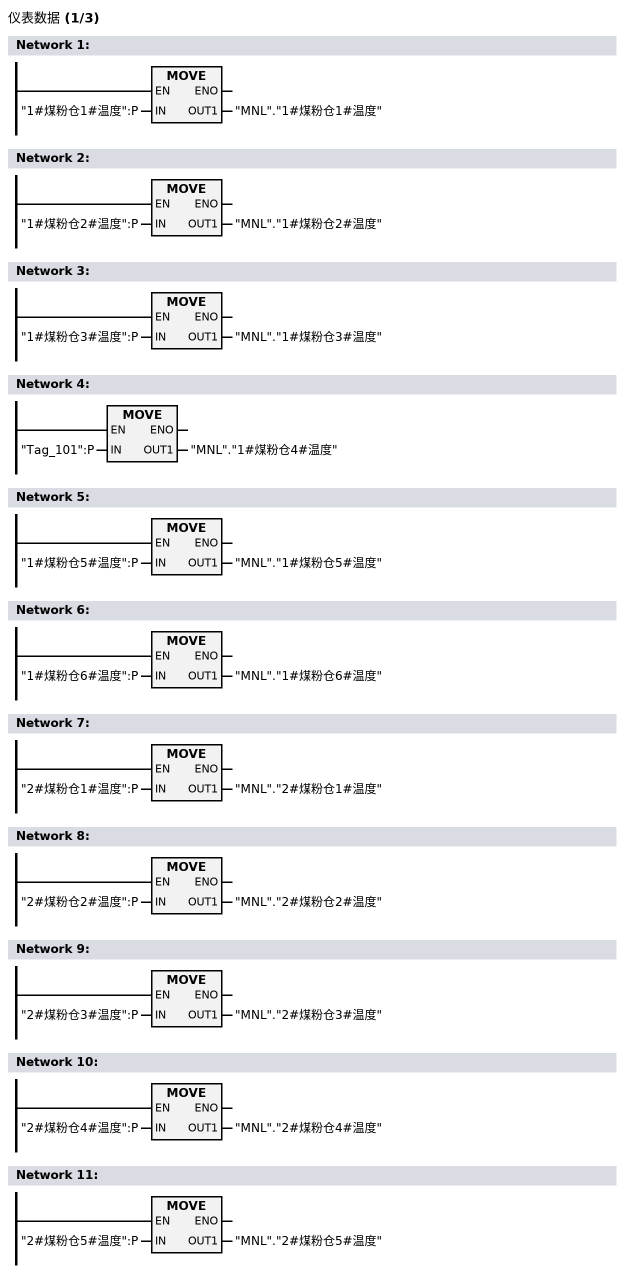
   RUNG wire#powerrail
      { S7_GenerateENO := "TRUE" } Move(in := "1#煤粉仓1#温度":P, out1 => "MNL"."1#煤粉仓1#温度")
   END_RUNG
   // the same network as SCL:
   "MNL"."1#煤粉仓1#温度" := "1#煤粉仓1#温度":P;
END_REGION
